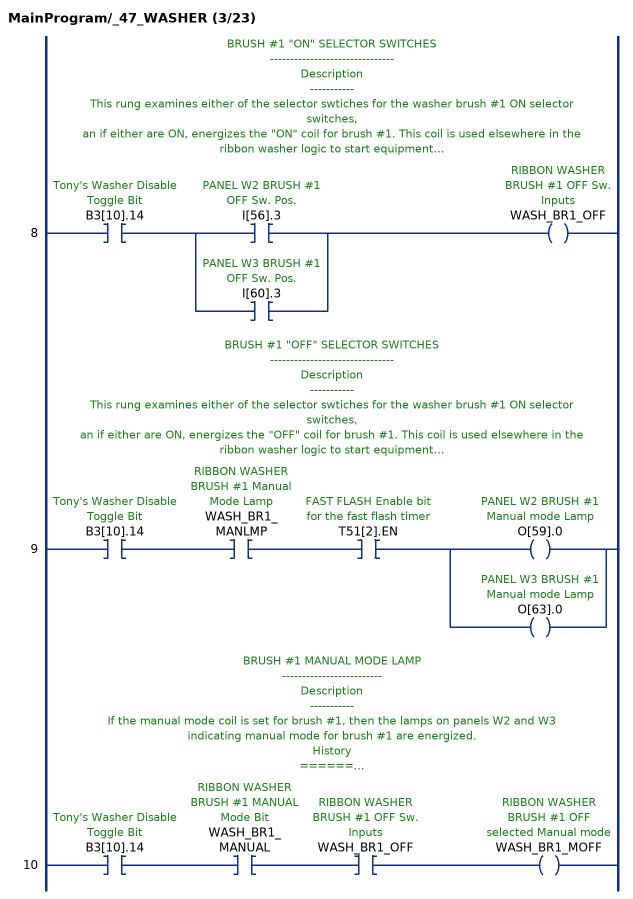
   // BRUSH #1 "ON" SELECTOR SWITCHES
   // -------------------------------
   // Description
   // -----------
   // This rung examines either of the selector swtiches for the washer brush #1 ON selector switches,
   // an if either are ON, energizes the "ON" coil for brush #1. This coil is used elsewhere in the
   // ribbon washer logic to start equipment.
   // History
   // =======
   // DATE        DESCRIPTION                                              PROGRAMMER
   // ----        -----------                                              ----------
   // 1/29/96     Entered rung and coil comments.                          WAS
   8: XIC(B3[10].14)[XIC(I[56].3) ,XIC(I[60].3) ]OTE(WASH_BR1_OFF);
   // BRUSH #1 "OFF" SELECTOR SWITCHES
   // -------------------------------
   // Description
   // -----------
   // This rung examines either of the selector swtiches for the washer brush #1 ON selector switches,
   // an if either are ON, energizes the "OFF" coil for brush #1. This coil is used elsewhere in the
   // ribbon washer logic to start equipment.
   // History
   // =======
   // DATE        DESCRIPTION                                              PROGRAMMER
   // ----        -----------                                              ----------
   // 1/29/96     Entered rung and coil comments.                          WAS
   9: XIC(B3[10].14)XIC(WASH_BR1_MANLMP)XIC(T51[2].EN)[OTE(O[59].0) ,OTE(O[63].0) ];
   // BRUSH #1 MANUAL MODE LAMP
   // -------------------------
   // Description
   // -----------
   // If the manual mode coil is set for brush #1, then the lamps on panels W2 and W3
   // indicating manual mode for brush #1 are energized.
   // History
   // =======
   // DATE        DESCRIPTION                                              PROGRAMMER
   // ----        -----------                                              ----------
   // 1/29/96     Entered rung and coil comments.                          WAS
   10: XIC(B3[10].14)XIC(WASH_BR1_MANUAL)XIC(WASH_BR1_OFF)OTE(WASH_BR1_MOFF);
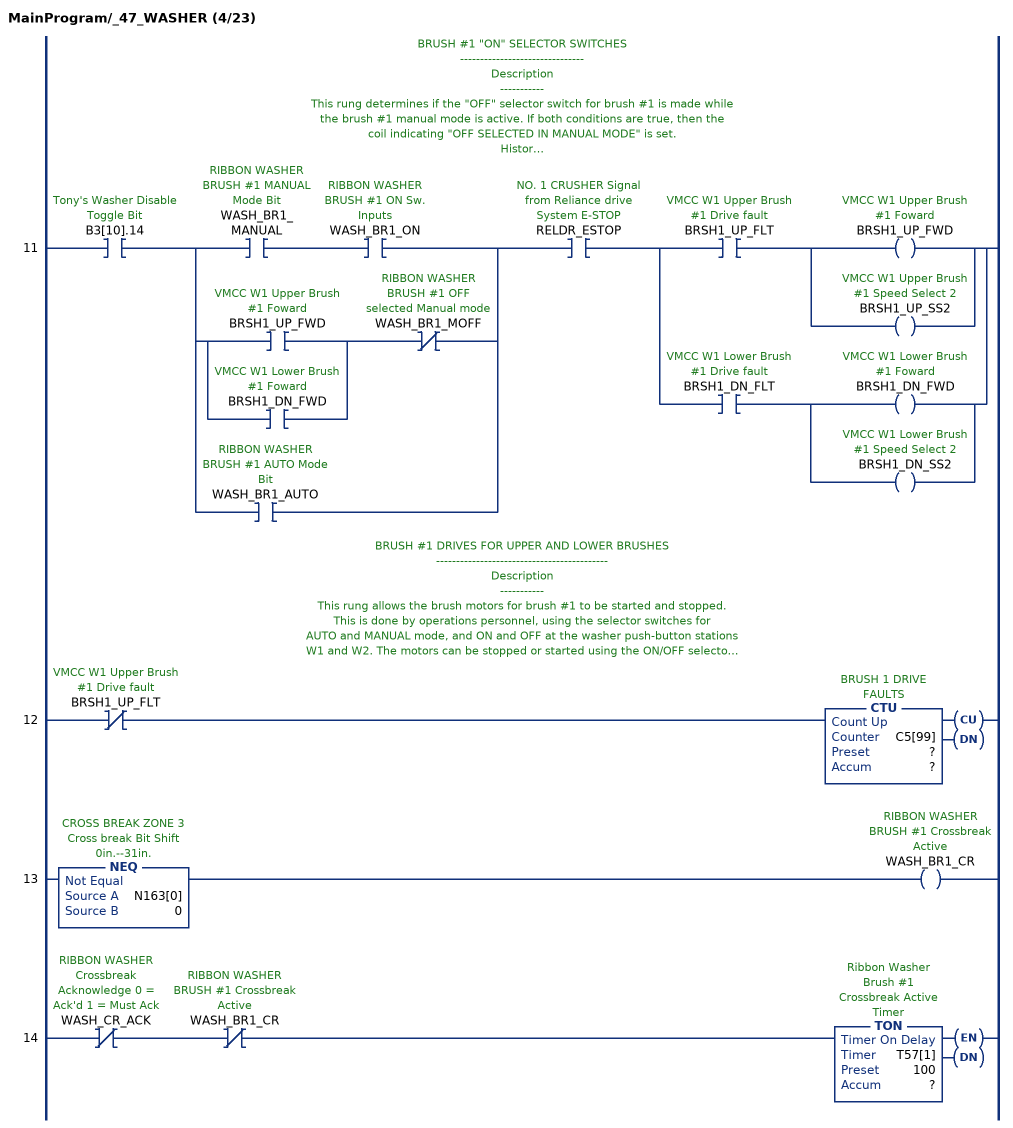
   // BRUSH #1 "ON" SELECTOR SWITCHES
   // -------------------------------
   // Description
   // -----------
   // This rung determines if the "OFF" selector switch for brush #1 is made while
   // the brush #1 manual mode is active. If both conditions are true, then the
   // coil indicating "OFF SELECTED IN MANUAL MODE" is set.
   // History
   // =======
   // DATE        DESCRIPTION                                              PROGRAMMER
   // ----        -----------                                              ----------
   // 1/29/96     Entered rung and coil comments.                          WAS
   11: XIC(B3[10].14)[XIC(WASH_BR1_MANUAL) XIC(WASH_BR1_ON) ,[XIC(BRSH1_UP_FWD) ,XIC(BRSH1_DN_FWD) ] XIO(WASH_BR1_MOFF) ,XIC(WASH_BR1_AUTO) ]XIC(RELDR_ESTOP)[XIC(BRSH1_UP_FLT) [OTE(BRSH1_UP_FWD) ,OTE(BRSH1_UP_SS2) ] ,XIC(BRSH1_DN_FLT) [OTE(BRSH1_DN_FWD) ,OTE(BRSH1_DN_SS2) ] ];
   // BRUSH #1 DRIVES FOR UPPER AND LOWER BRUSHES
   // -------------------------------------------
   // Description
   // -----------
   // This rung allows the brush motors for brush #1 to be started and stopped.
   // This is done by operations personnel, using the selector switches for
   // AUTO and MANUAL mode, and ON and OFF at the washer push-button stations
   // W1 and W2. The motors can be stopped or started using the ON/OFF selector
   // switch if and only if the washer is in manual mode.
   // History
   // =======
   // DATE        DESCRIPTION                                              PROGRAMMER
   // ----        -----------                                              ----------
   // 1/29/96     Entered rung and coil comments.                          WAS
   12: XIO(BRSH1_UP_FLT)CTU(C5[99],?,?);
   13: NEQ(N163[0],0)OTE(WASH_BR1_CR);
   14: XIO(WASH_CR_ACK)XIO(WASH_BR1_CR)TON(T57[1],?,?);
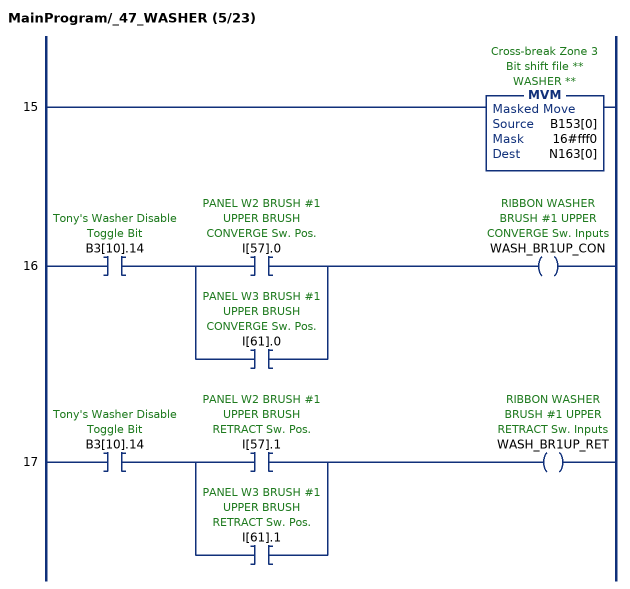
   15: MVM(B153[0],16#fff0,N163[0]);
   16: XIC(B3[10].14)[XIC(I[57].0) ,XIC(I[61].0) ]OTE(WASH_BR1UP_CON);
   17: XIC(B3[10].14)[XIC(I[57].1) ,XIC(I[61].1) ]OTE(WASH_BR1UP_RET);
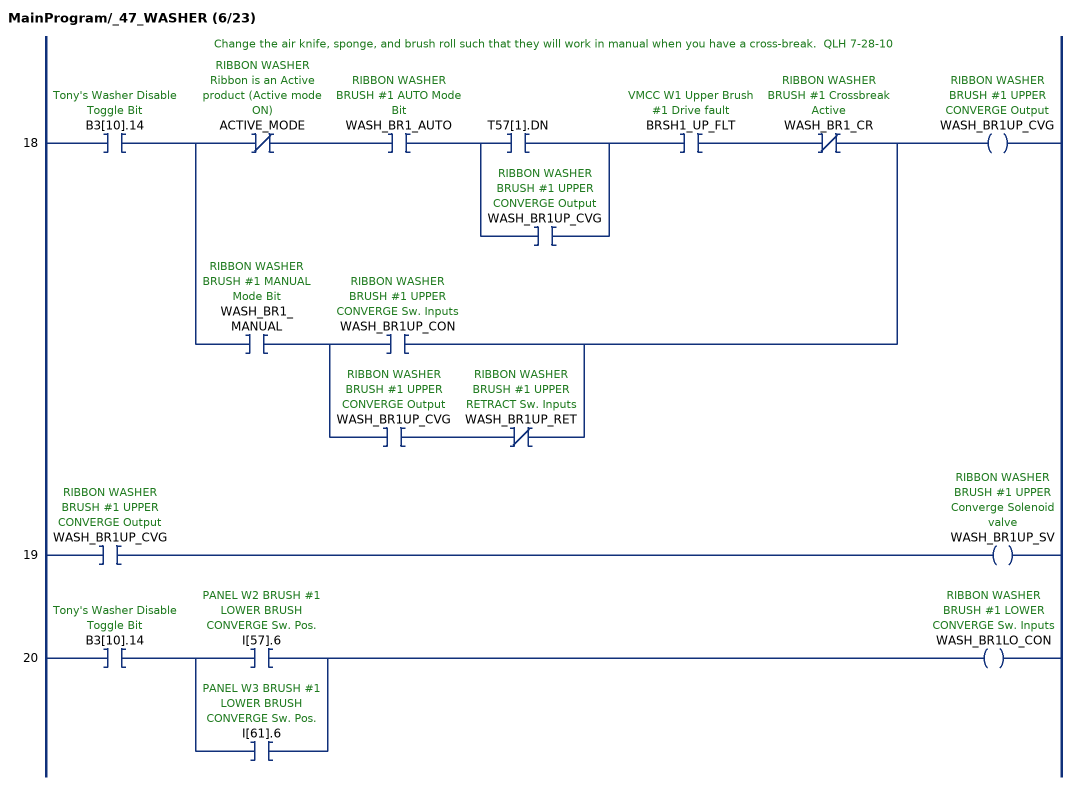
   // Change the air knife, sponge, and brush roll such that they will work in manual when you have a cross-break.  QLH 7-28-10
   18: XIC(B3[10].14)[XIO(ACTIVE_MODE) XIC(WASH_BR1_AUTO) [XIC(T57[1].DN) ,XIC(WASH_BR1UP_CVG) ] XIC(BRSH1_UP_FLT) XIO(WASH_BR1_CR) ,XIC(WASH_BR1_MANUAL) [XIC(WASH_BR1UP_CON) ,XIC(WASH_BR1UP_CVG) XIO(WASH_BR1UP_RET) ] ]OTE(WASH_BR1UP_CVG);
   19: XIC(WASH_BR1UP_CVG)OTE(WASH_BR1UP_SV);
   20: XIC(B3[10].14)[XIC(I[57].6) ,XIC(I[61].6) ]OTE(WASH_BR1LO_CON);
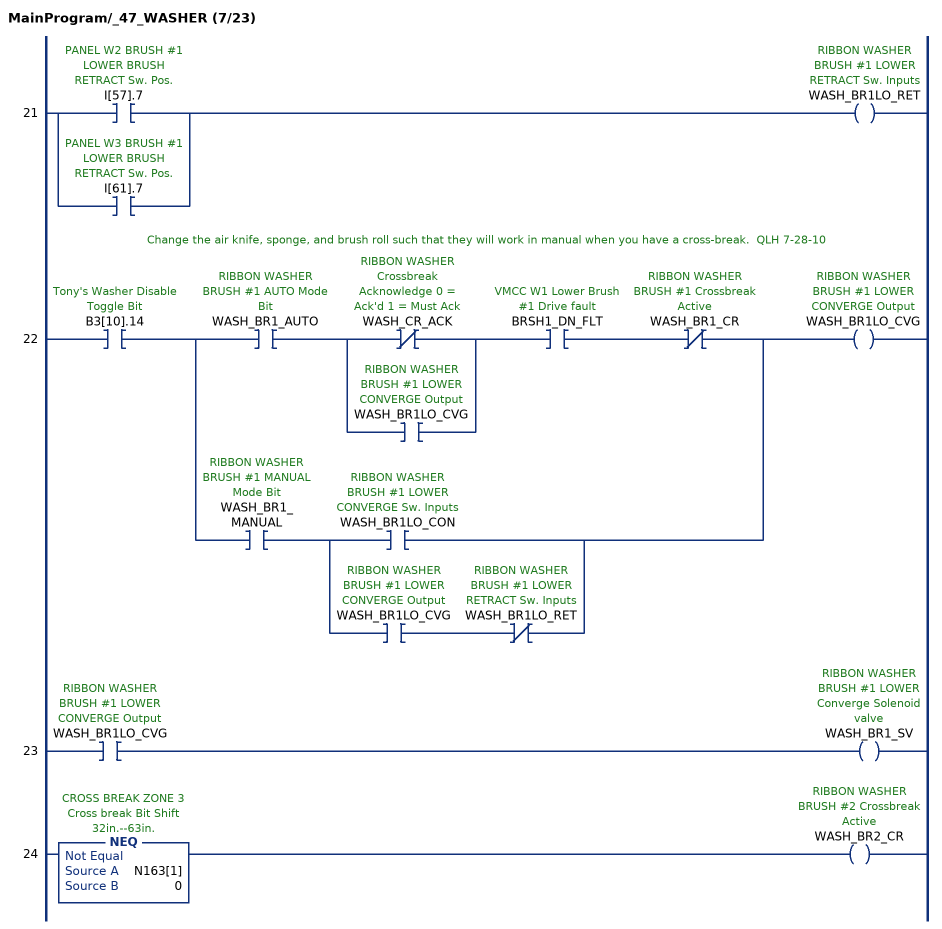
   21: [XIC(I[57].7) ,XIC(I[61].7) ]OTE(WASH_BR1LO_RET);
   // Change the air knife, sponge, and brush roll such that they will work in manual when you have a cross-break.  QLH 7-28-10
   22: XIC(B3[10].14)[XIC(WASH_BR1_AUTO) [XIO(WASH_CR_ACK) ,XIC(WASH_BR1LO_CVG) ] XIC(BRSH1_DN_FLT) XIO(WASH_BR1_CR) ,XIC(WASH_BR1_MANUAL) [XIC(WASH_BR1LO_CON) ,XIC(WASH_BR1LO_CVG) XIO(WASH_BR1LO_RET) ] ]OTE(WASH_BR1LO_CVG);
   23: XIC(WASH_BR1LO_CVG)OTE(WASH_BR1_SV);
   24: NEQ(N163[1],0)OTE(WASH_BR2_CR);
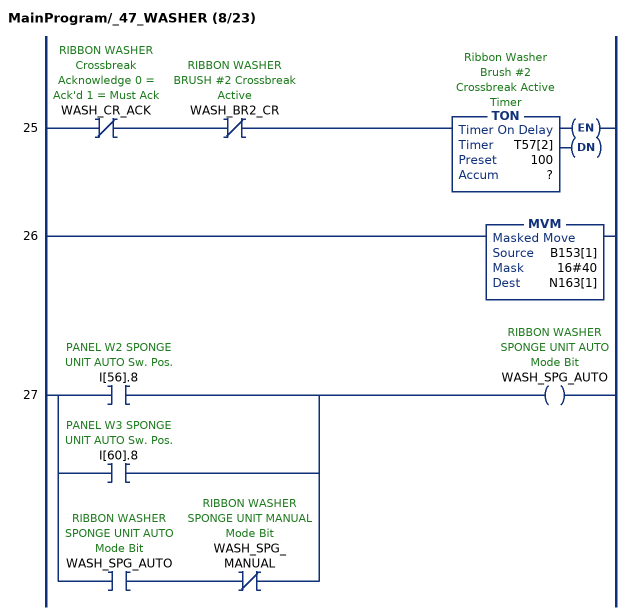
   25: XIO(WASH_CR_ACK)XIO(WASH_BR2_CR)TON(T57[2],?,?);
   26: MVM(B153[1],16#40,N163[1]);
   27: [[XIC(I[56].8) ,XIC(I[60].8) ] ,XIC(WASH_SPG_AUTO) XIO(WASH_SPG_MANUAL) ]OTE(WASH_SPG_AUTO);
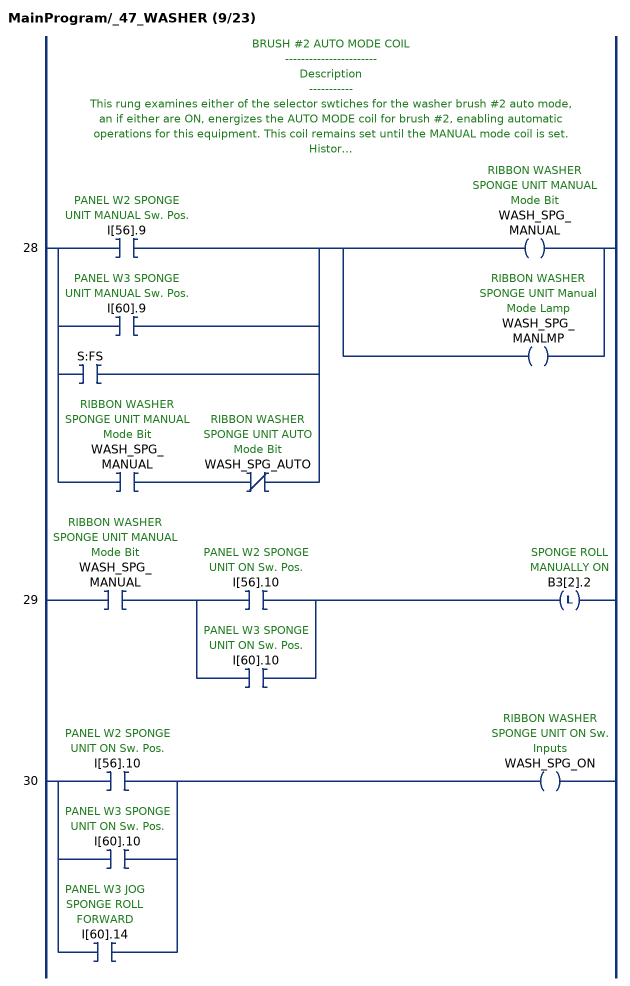
   // BRUSH #2 AUTO MODE COIL
   // -----------------------
   // Description
   // -----------
   // This rung examines either of the selector swtiches for the washer brush #2 auto mode,
   // an if either are ON, energizes the AUTO MODE coil for brush #2, enabling automatic
   // operations for this equipment. This coil remains set until the MANUAL mode coil is set.
   // History
   // =======
   // DATE        DESCRIPTION                                              PROGRAMMER
   // ----        -----------                                              ----------
   // 1/29/96     Entered rung and coil comments.                          WAS
   28: [[XIC(I[56].9) ,XIC(I[60].9) ,XIC(S:FS) ] ,XIC(WASH_SPG_MANUAL) XIO(WASH_SPG_AUTO) ][OTE(WASH_SPG_MANUAL) ,OTE(WASH_SPG_MANLMP) ];
   29: XIC(WASH_SPG_MANUAL)[XIC(I[56].10) ,XIC(I[60].10) ]OTL(B3[2].2);
   30: [XIC(I[56].10) ,XIC(I[60].10) ,XIC(I[60].14) ]OTE(WASH_SPG_ON);
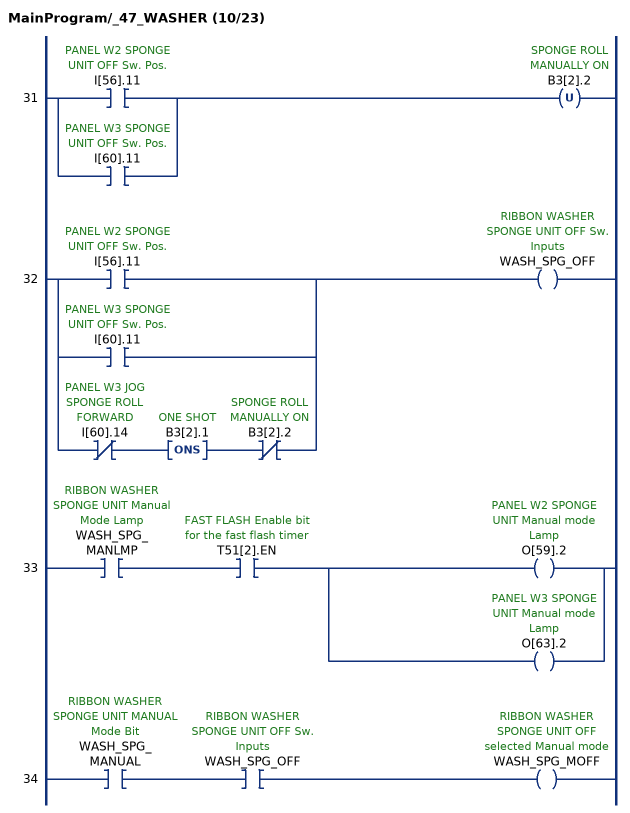
   31: [XIC(I[56].11) ,XIC(I[60].11) ]OTU(B3[2].2);
   32: [XIC(I[56].11) ,XIC(I[60].11) ,XIO(I[60].14) ONS(B3[2].1) XIO(B3[2].2) ]OTE(WASH_SPG_OFF);
   33: XIC(WASH_SPG_MANLMP)XIC(T51[2].EN)[OTE(O[59].2) ,OTE(O[63].2) ];
   34: XIC(WASH_SPG_MANUAL)XIC(WASH_SPG_OFF)OTE(WASH_SPG_MOFF);
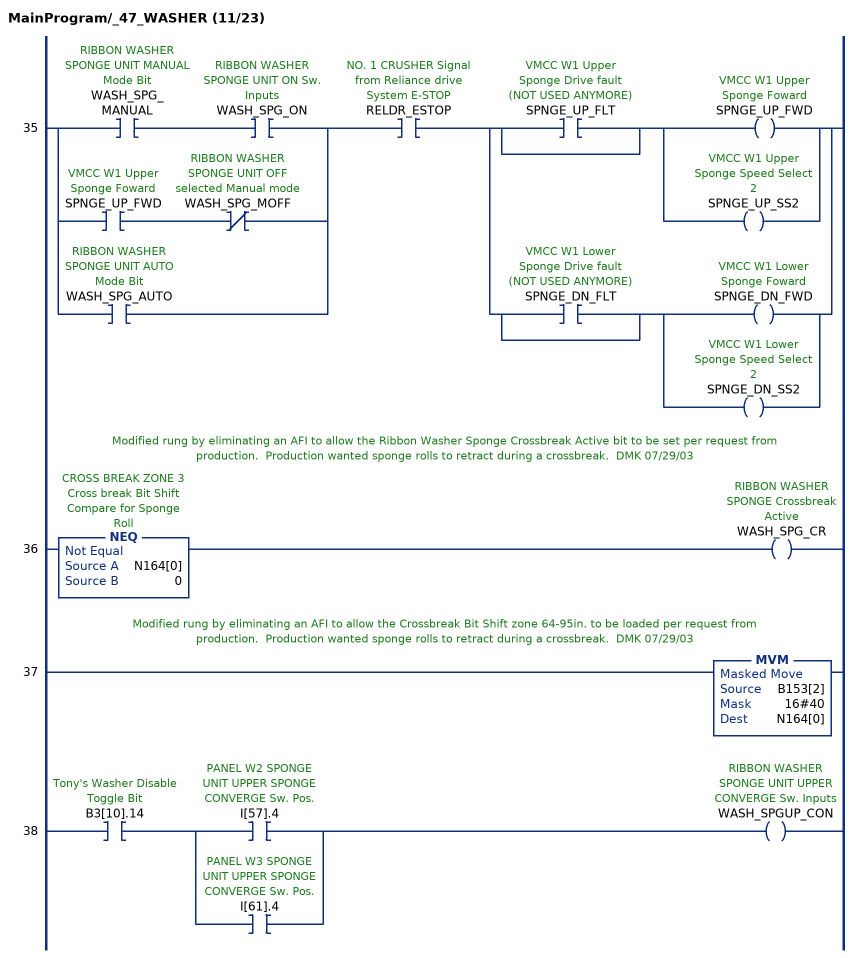
   35: [XIC(WASH_SPG_MANUAL) XIC(WASH_SPG_ON) ,XIC(SPNGE_UP_FWD) XIO(WASH_SPG_MOFF) ,XIC(WASH_SPG_AUTO) ]XIC(RELDR_ESTOP)[[XIC(SPNGE_UP_FLT) ,] [OTE(SPNGE_UP_FWD) ,OTE(SPNGE_UP_SS2) ] ,[XIC(SPNGE_DN_FLT) ,] [OTE(SPNGE_DN_FWD) ,OTE(SPNGE_DN_SS2) ] ];
   // Modified rung by eliminating an AFI to allow the Ribbon Washer Sponge Crossbreak Active bit to be set per request from
   // production.  Production wanted sponge rolls to retract during a crossbreak.  DMK 07/29/03
   36: NEQ(N164[0],0)OTE(WASH_SPG_CR);
   // Modified rung by eliminating an AFI to allow the Crossbreak Bit Shift zone 64-95in. to be loaded per request from
   // production.  Production wanted sponge rolls to retract during a crossbreak.  DMK 07/29/03
   37: MVM(B153[2],16#40,N164[0]);
   38: XIC(B3[10].14)[XIC(I[57].4) ,XIC(I[61].4) ]OTE(WASH_SPGUP_CON);
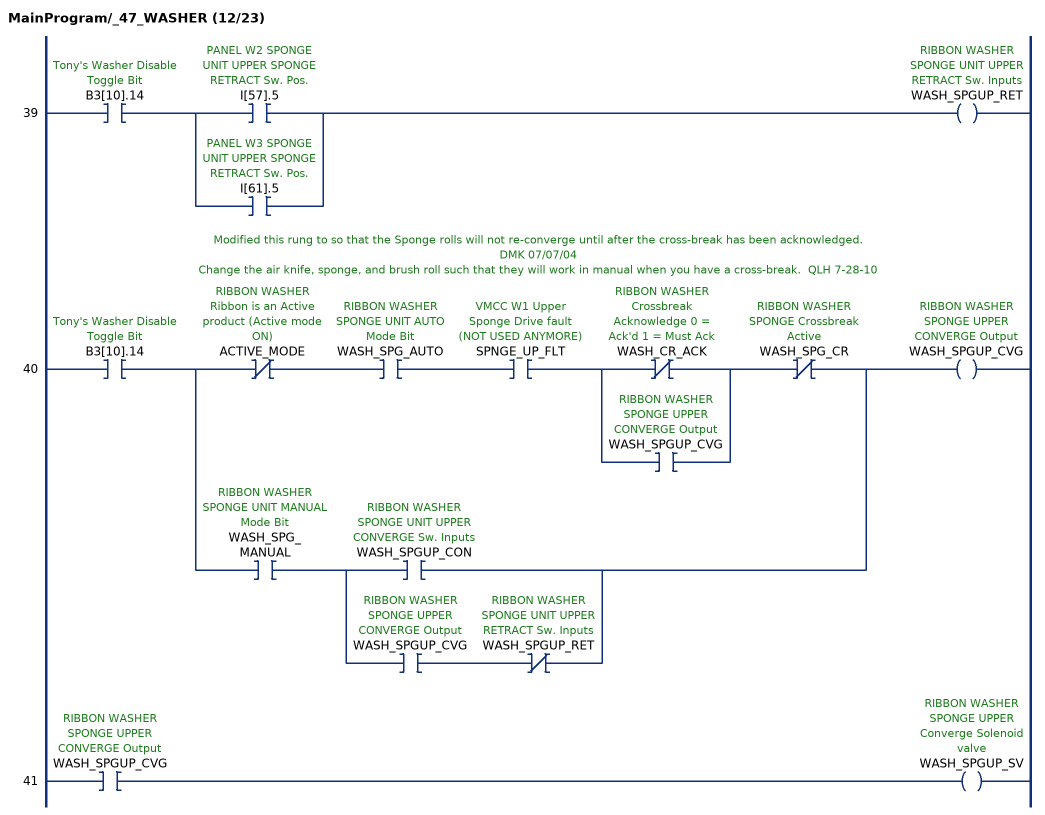
   39: XIC(B3[10].14)[XIC(I[57].5) ,XIC(I[61].5) ]OTE(WASH_SPGUP_RET);
   // Modified this rung to so that the Sponge rolls will not re-converge until after the cross-break has been acknowledged.
   // DMK 07/07/04
   // Change the air knife, sponge, and brush roll such that they will work in manual when you have a cross-break.  QLH 7-28-10
   40: XIC(B3[10].14)[XIO(ACTIVE_MODE) XIC(WASH_SPG_AUTO) XIC(SPNGE_UP_FLT) [XIO(WASH_CR_ACK) ,XIC(WASH_SPGUP_CVG) ] XIO(WASH_SPG_CR) ,XIC(WASH_SPG_MANUAL) [XIC(WASH_SPGUP_CON) ,XIC(WASH_SPGUP_CVG) XIO(WASH_SPGUP_RET) ] ]OTE(WASH_SPGUP_CVG);
   41: XIC(WASH_SPGUP_CVG)OTE(WASH_SPGUP_SV);
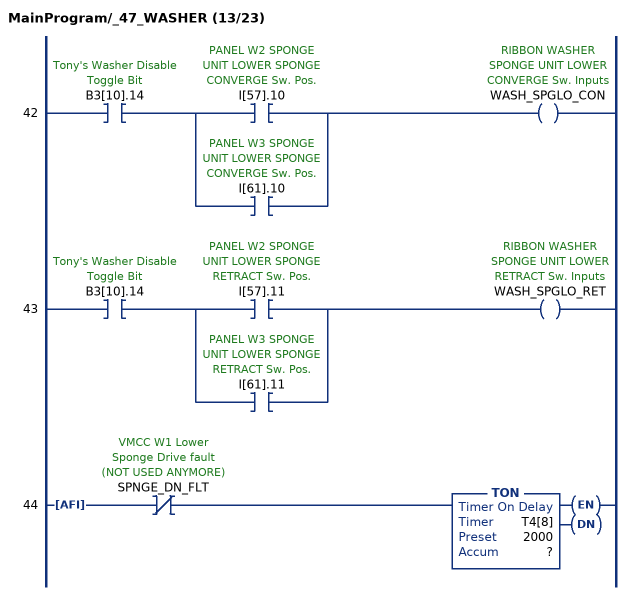
   42: XIC(B3[10].14)[XIC(I[57].10) ,XIC(I[61].10) ]OTE(WASH_SPGLO_CON);
   43: XIC(B3[10].14)[XIC(I[57].11) ,XIC(I[61].11) ]OTE(WASH_SPGLO_RET);
   44: AFI()XIO(SPNGE_DN_FLT)TON(T4[8],?,?);
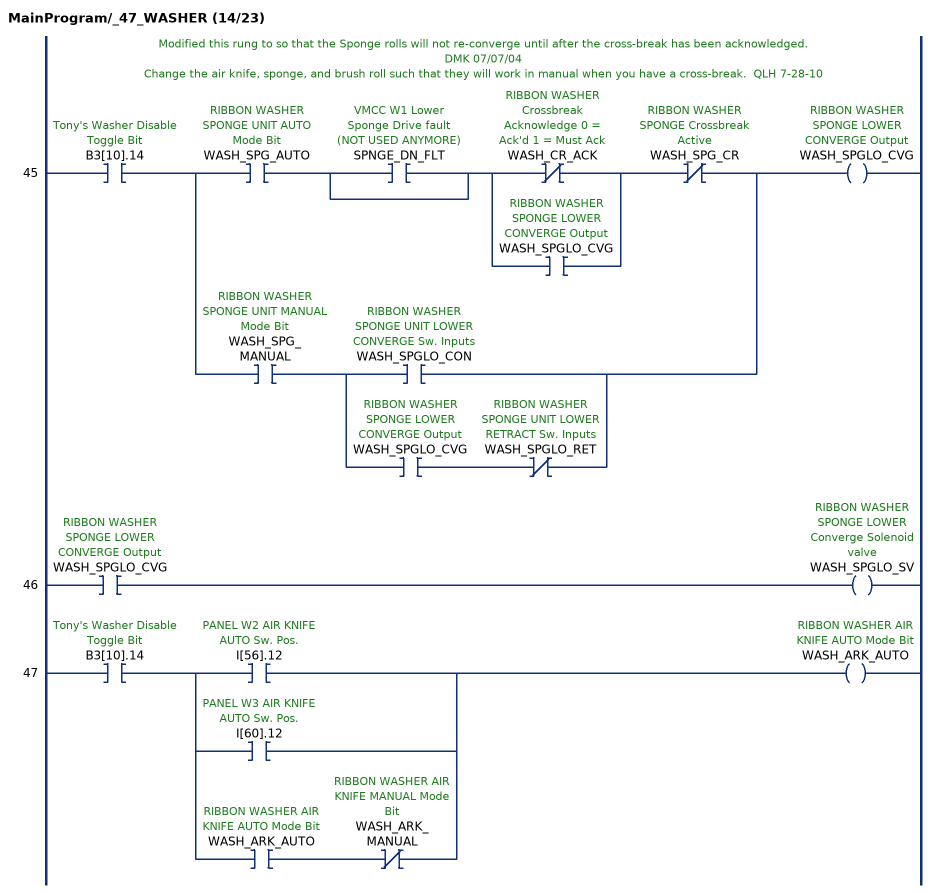
   // Modified this rung to so that the Sponge rolls will not re-converge until after the cross-break has been acknowledged.
   // DMK 07/07/04
   // Change the air knife, sponge, and brush roll such that they will work in manual when you have a cross-break.  QLH 7-28-10
   45: XIC(B3[10].14)[XIC(WASH_SPG_AUTO) [XIC(SPNGE_DN_FLT) ,] [XIO(WASH_CR_ACK) ,XIC(WASH_SPGLO_CVG) ] XIO(WASH_SPG_CR) ,XIC(WASH_SPG_MANUAL) [XIC(WASH_SPGLO_CON) ,XIC(WASH_SPGLO_CVG) XIO(WASH_SPGLO_RET) ] ]OTE(WASH_SPGLO_CVG);
   46: XIC(WASH_SPGLO_CVG)OTE(WASH_SPGLO_SV);
   47: XIC(B3[10].14)[[XIC(I[56].12) ,XIC(I[60].12) ] ,XIC(WASH_ARK_AUTO) XIO(WASH_ARK_MANUAL) ]OTE(WASH_ARK_AUTO);
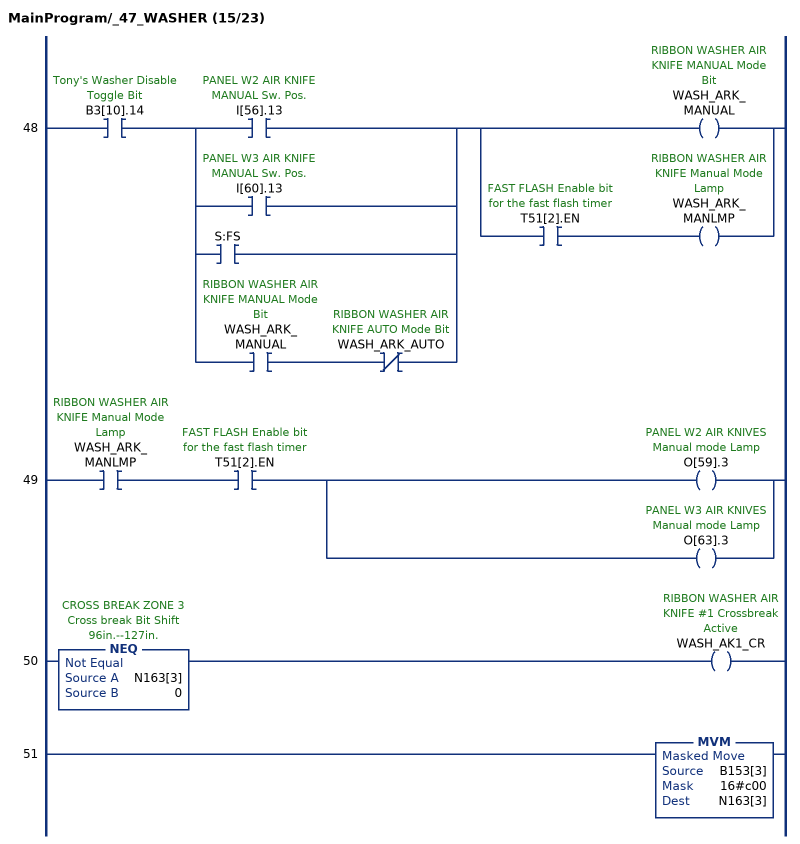
   48: XIC(B3[10].14)[[XIC(I[56].13) ,XIC(I[60].13) ,XIC(S:FS) ] ,XIC(WASH_ARK_MANUAL) XIO(WASH_ARK_AUTO) ][OTE(WASH_ARK_MANUAL) ,XIC(T51[2].EN) OTE(WASH_ARK_MANLMP) ];
   49: XIC(WASH_ARK_MANLMP)XIC(T51[2].EN)[OTE(O[59].3) ,OTE(O[63].3) ];
   50: NEQ(N163[3],0)OTE(WASH_AK1_CR);
   51: MVM(B153[3],16#c00,N163[3]);
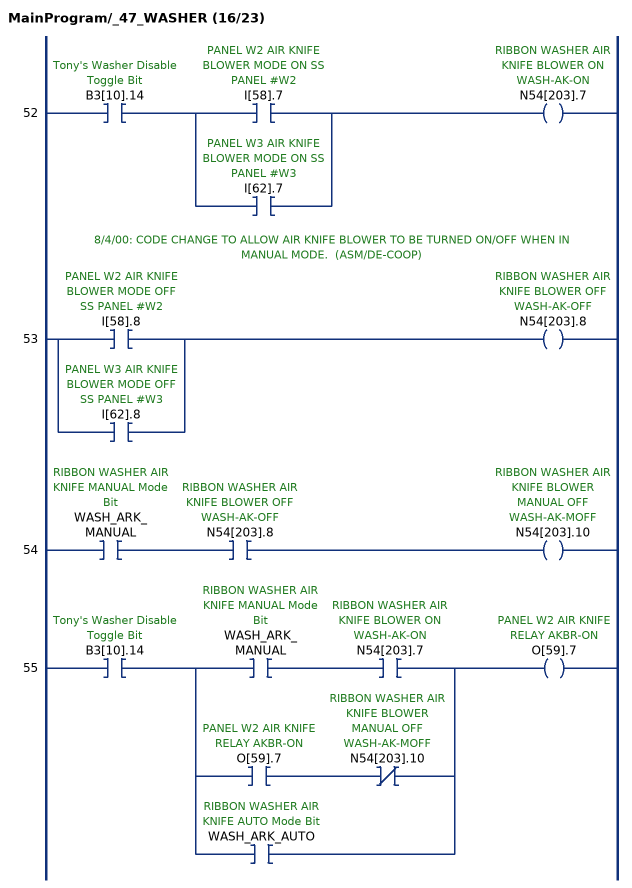
   52: XIC(B3[10].14)[XIC(I[58].7) ,XIC(I[62].7) ]OTE(N54[203].7);
   // 8/4/00: CODE CHANGE TO ALLOW AIR KNIFE BLOWER TO BE TURNED ON/OFF WHEN IN MANUAL MODE.  (ASM/DE-COOP)
   53: [XIC(I[58].8) ,XIC(I[62].8) ]OTE(N54[203].8);
   54: XIC(WASH_ARK_MANUAL)XIC(N54[203].8)OTE(N54[203].10);
   55: XIC(B3[10].14)[[XIC(WASH_ARK_MANUAL) XIC(N54[203].7) ,XIC(O[59].7) XIO(N54[203].10) ] ,XIC(WASH_ARK_AUTO) ]OTE(O[59].7);
